// TIA Portal project "EbAndon v4_00_036" (V15) (continued)
   // pnText[239] := WSTRING#'//';
   // pnText[240] := WSTRING#'//';
   // pnText[241] := WSTRING#'//';
   // pnText[242] := WSTRING#'//';
   // pnText[243] := WSTRING#'//';
   // pnText[244] := WSTRING#'//';
   // pnText[245] := WSTRING#'//';
   // pnText[246] := WSTRING#'//';
   // pnText[247] := WSTRING#'//';
   // pnText[248] := WSTRING#'//';
   // pnText[249] := WSTRING#'//';
   // pnText[250] := WSTRING#'//';
   // pnText[251] := WSTRING#'//';
   // pnText[252] := WSTRING#'//';
   // pnText[253] := WSTRING#'//';
   // pnText[254] := WSTRING#'//';
   // pnText[255] := WSTRING#'//';
   // pnText[256] := WSTRING#'//';
   // pnText[257] := WSTRING#'//';
   // pnText[258] := WSTRING#'//';
   // pnText[259] := WSTRING#'//';
   // pnText[260] := WSTRING#'//';
   // pnText[261] := WSTRING#'//';
   // pnText[262] := WSTRING#'//';
   // pnText[263] := WSTRING#'//';
   // pnText[264] := WSTRING#'//';
   // pnText[265] := WSTRING#'//';
   // pnText[266] := WSTRING#'//';
   // pnText[267] := WSTRING#'//';
   // pnText[268] := WSTRING#'//';
   // pnText[269] := WSTRING#'//';
   // pnText[270] := WSTRING#'//';
   // pnText[271] := WSTRING#'//';
   // pnText[272] := WSTRING#'//';
   // pnText[273] := WSTRING#'//';
   // pnText[274] := WSTRING#'//';
   // pnText[275] := WSTRING#'//';
   // pnText[276] := WSTRING#'//';
   // pnText[277] := WSTRING#'//';
   // pnText[278] := WSTRING#'//';
   // pnText[279] := WSTRING#'//';
   // pnText[280] := WSTRING#'//';
   // pnText[281] := WSTRING#'//';
   // pnText[282] := WSTRING#'//';
   // pnText[283] := WSTRING#'//';
   // pnText[284] := WSTRING#'//';
   // pnText[285] := WSTRING#'//';
   // pnText[286] := WSTRING#'//';
   // pnText[287] := WSTRING#'//';
   // pnText[288] := WSTRING#'//';
   // pnText[289] := WSTRING#'//';
   // pnText[290] := WSTRING#'//';
   // pnText[291] := WSTRING#'//';
   // pnText[292] := WSTRING#'//';
   // pnText[293] := WSTRING#'//';
   // pnText[294] := WSTRING#'//';
   // pnText[295] := WSTRING#'//';
   // pnText[296] := WSTRING#'//';
   // pnText[297] := WSTRING#'//';
   // pnText[298] := WSTRING#'//';
   // pnText[299] := WSTRING#'//';
   // pnText[300] := WSTRING#'//';
   // pnText[301] := WSTRING#'//';
   // pnText[302] := WSTRING#'//';
   // pnText[303] := WSTRING#'//';
   // pnText[304] := WSTRING#'//';
   // pnText[305] := WSTRING#'//';
   // pnText[306] := WSTRING#'//';
   // pnText[307] := WSTRING#'//';
   // pnText[308] := WSTRING#'//';
   // pnText[309] := WSTRING#'//';
   // pnText[310] := WSTRING#'//';
   // pnText[311] := WSTRING#'//';
   // pnText[312] := WSTRING#'//';
   // pnText[313] := WSTRING#'//';
   // pnText[314] := WSTRING#'//';
   // pnText[315] := WSTRING#'//';
   // pnText[316] := WSTRING#'//';
   // pnText[317] := WSTRING#'//';
   // pnText[318] := WSTRING#'//';
   // pnText[319] := WSTRING#'//';
   // pnText[320] := WSTRING#'//';
   // pnText[321] := WSTRING#'//';
   // pnText[322] := WSTRING#'//';
   // pnText[323] := WSTRING#'//';
   // pnText[324] := WSTRING#'//';
   // pnText[325] := WSTRING#'//';
   // pnText[326] := WSTRING#'//';
   // pnText[327] := WSTRING#'//';
   // pnText[328] := WSTRING#'//';
   // pnText[329] := WSTRING#'//';
   // pnText[330] := WSTRING#'//';
   // pnText[331] := WSTRING#'//';
   // pnText[332] := WSTRING#'//';
   // pnText[333] := WSTRING#'//';
   // pnText[334] := WSTRING#'//';
   // pnText[335] := WSTRING#'//';
   // pnText[336] := WSTRING#'//';
   // pnText[337] := WSTRING#'//';
   // pnText[338] := WSTRING#'//';
   // pnText[339] := WSTRING#'//';
   // pnText[340] := WSTRING#'//';
   // pnText[341] := WSTRING#'//';
   // pnText[342] := WSTRING#'//';
   // pnText[343] := WSTRING#'//';
   // pnText[344] := WSTRING#'//';
   // pnText[345] := WSTRING#'//';
   // pnText[346] := WSTRING#'//';
   // pnText[347] := WSTRING#'//';
   // pnText[348] := WSTRING#'//';
   // pnText[349] := WSTRING#'//';
   // pnText[350] := WSTRING#'//';
   // pnText[351] := WSTRING#'//';
   // pnText[352] := WSTRING#'//';
   // pnText[353] := WSTRING#'//';
   // pnText[354] := WSTRING#'//';
   // pnText[355] := WSTRING#'//';
   // pnText[356] := WSTRING#'//';
   // pnText[357] := WSTRING#'//';
   // pnText[358] := WSTRING#'//';
   // pnText[359] := WSTRING#'//';
   // pnText[360] := WSTRING#'//';
   // pnText[361] := WSTRING#'//';
   // pnText[362] := WSTRING#'//';
   // pnText[363] := WSTRING#'//';
   // pnText[364] := WSTRING#'//';
   // pnText[365] := WSTRING#'//';
   // pnText[366] := WSTRING#'//';
   // pnText[367] := WSTRING#'//';
   // pnText[368] := WSTRING#'//';
   // pnText[369] := WSTRING#'//';
   // pnText[370] := WSTRING#'//';
   // pnText[371] := WSTRING#'//';
   // pnText[372] := WSTRING#'//';
   // pnText[373] := WSTRING#'//';
   // pnText[374] := WSTRING#'//';
   // pnText[375] := WSTRING#'//';
   // pnText[376] := WSTRING#'//';
   // pnText[377] := WSTRING#'//';
   // pnText[378] := WSTRING#'//';
   // pnText[379] := WSTRING#'//';
   // pnText[380] := WSTRING#'//';
   // pnText[381] := WSTRING#'//';
   // pnText[382] := WSTRING#'//';
   // pnText[383] := WSTRING#'//';
   // pnText[384] := WSTRING#'//';
   // pnText[385] := WSTRING#'//';
   // pnText[386] := WSTRING#'//';
   // pnText[387] := WSTRING#'//';
   // pnText[388] := WSTRING#'//';
   // pnText[389] := WSTRING#'//';
   // pnText[390] := WSTRING#'//';
   // pnText[391] := WSTRING#'//';
   // pnText[392] := WSTRING#'//';
   // pnText[393] := WSTRING#'//';
   // pnText[394] := WSTRING#'//';
   // pnText[395] := WSTRING#'//';
   // pnText[396] := WSTRING#'//';
   // pnText[397] := WSTRING#'//';
   // pnText[398] := WSTRING#'//';
   // pnText[399] := WSTRING#'//';
   // pnText[400] := WSTRING#'//';
   // pnText[401] := WSTRING#'//';
   // pnText[402] := WSTRING#'//';
   // pnText[403] := WSTRING#'//';
   // pnText[404] := WSTRING#'//';
   // pnText[405] := WSTRING#'//';
   // pnText[406] := WSTRING#'//';
   // pnText[407] := WSTRING#'//';
   // pnText[408] := WSTRING#'//';
   // pnText[409] := WSTRING#'//';
   // pnText[410] := WSTRING#'//';
   // pnText[411] := WSTRING#'//';
   // pnText[412] := WSTRING#'//';
   // pnText[413] := WSTRING#'//';
   // pnText[414] := WSTRING#'//';
   // pnText[415] := WSTRING#'//';
   // pnText[416] := WSTRING#'//';
   // pnText[417] := WSTRING#'//';
   // pnText[418] := WSTRING#'//';
   // pnText[419] := WSTRING#'//';
   // pnText[420] := WSTRING#'//';
   // pnText[421] := WSTRING#'//';
   // pnText[422] := WSTRING#'//';
   // pnText[423] := WSTRING#'//';
   // pnText[424] := WSTRING#'//';
   // pnText[425] := WSTRING#'//';
   // pnText[426] := WSTRING#'//';
   // pnText[427] := WSTRING#'//';
   // pnText[428] := WSTRING#'//';
   // pnText[429] := WSTRING#'//';
   // pnText[430] := WSTRING#'//';
   // pnText[431] := WSTRING#'//';
   // pnText[432] := WSTRING#'//';
   // pnText[433] := WSTRING#'//';
   // pnText[434] := WSTRING#'//';
   // pnText[435] := WSTRING#'//';
   // pnText[436] := WSTRING#'//';
   // pnText[437] := WSTRING#'//';
   // pnText[438] := WSTRING#'//';
   // pnText[439] := WSTRING#'//';
   // pnText[440] := WSTRING#'//';
   // pnText[441] := WSTRING#'//';
   // pnText[442] := WSTRING#'//';
   // pnText[443] := WSTRING#'//';
   // pnText[444] := WSTRING#'//';
   // pnText[445] := WSTRING#'//';
   // pnText[446] := WSTRING#'//';
   // pnText[447] := WSTRING#'//';
   // pnText[448] := WSTRING#'//';
   // pnText[449] := WSTRING#'//';
   // pnText[450] := WSTRING#'//';
   // pnText[451] := WSTRING#'//';
   // pnText[452] := WSTRING#'//';
   // pnText[453] := WSTRING#'//';
   // pnText[454] := WSTRING#'//';
   // pnText[455] := WSTRING#'//';
   // pnText[456] := WSTRING#'//';
   // pnText[457] := WSTRING#'//';
   // pnText[458] := WSTRING#'//';
   // pnText[459] := WSTRING#'//';
   // pnText[460] := WSTRING#'//';
   // pnText[461] := WSTRING#'//';
   // pnText[462] := WSTRING#'//';
   // pnText[463] := WSTRING#'//';
   // pnText[464] := WSTRING#'//';
   // pnText[465] := WSTRING#'//';
   // pnText[466] := WSTRING#'//';
   // pnText[467] := WSTRING#'//';
   // pnText[468] := WSTRING#'//';
   // pnText[469] := WSTRING#'//';
   // pnText[470] := WSTRING#'//';
   // pnText[471] := WSTRING#'//';
   // pnText[472] := WSTRING#'//';
   // pnText[473] := WSTRING#'//';
   // pnText[474] := WSTRING#'//';
   // pnText[475] := WSTRING#'//';
   // pnText[476] := WSTRING#'//';
   // pnText[477] := WSTRING#'//';
   // pnText[478] := WSTRING#'//';
   // pnText[479] := WSTRING#'//';
   // pnText[480] := WSTRING#'//';
   // pnText[481] := WSTRING#'//';
   // pnText[482] := WSTRING#'//';
   // pnText[483] := WSTRING#'//';
   // pnText[484] := WSTRING#'//';
   // pnText[485] := WSTRING#'//';
   // pnText[486] := WSTRING#'//';
   // pnText[487] := WSTRING#'//';
   // pnText[488] := WSTRING#'//';
   // pnText[489] := WSTRING#'//';
   // pnText[490] := WSTRING#'//';
   // pnText[491] := WSTRING#'//';
   // pnText[492] := WSTRING#'//';
   // pnText[493] := WSTRING#'//';
   // pnText[494] := WSTRING#'//';
   // pnText[495] := WSTRING#'//';
   // pnText[496] := WSTRING#'//';
   // pnText[497] := WSTRING#'//';
   // pnText[498] := WSTRING#'//';
   // pnText[499] := WSTRING#'//';
   // pnText[500] := WSTRING#'//';
   // pnText[501] := WSTRING#'//';
   // pnText[502] := WSTRING#'//';
   // pnText[503] := WSTRING#'//';
   // pnText[504] := WSTRING#'//';
   // pnText[505] := WSTRING#'//';
   // pnText[506] := WSTRING#'//';
   // pnText[507] := WSTRING#'//';
   // pnText[508] := WSTRING#'//';
   // pnText[509] := WSTRING#'//';
   // pnText[510] := WSTRING#'//';
   // pnText[511] := WSTRING#'//';
   // pnText[512] := WSTRING#'//';
   // pnText[513] := WSTRING#'//';
   // pnText[514] := WSTRING#'//';
   // pnText[515] := WSTRING#'//';
   // pnText[516] := WSTRING#'//';
   // pnText[517] := WSTRING#'//';
   // pnText[518] := WSTRING#'//';
   // pnText[519] := WSTRING#'//';
   // pnText[520] := WSTRING#'//';
   // pnText[521] := WSTRING#'//';
   // pnText[522] := WSTRING#'//';
   // pnText[523] := WSTRING#'//';
   // pnText[524] := WSTRING#'//';
   // pnText[525] := WSTRING#'//';
   // pnText[526] := WSTRING#'//';
   // pnText[527] := WSTRING#'//';
   // pnText[528] := WSTRING#'//';
   // pnText[529] := WSTRING#'//';
   // pnText[530] := WSTRING#'//';
   // pnText[531] := WSTRING#'//';
   // pnText[532] := WSTRING#'//';
   // pnText[533] := WSTRING#'//';
   // pnText[534] := WSTRING#'//';
   // pnText[535] := WSTRING#'//';
   // pnText[536] := WSTRING#'//';
   // pnText[537] := WSTRING#'//';
   // pnText[538] := WSTRING#'//';
   // pnText[539] := WSTRING#'//';
   // pnText[540] := WSTRING#'//';
   // pnText[541] := WSTRING#'//';
   // pnText[542] := WSTRING#'//';
   // pnText[543] := WSTRING#'//';
   // pnText[544] := WSTRING#'//';
   // pnText[545] := WSTRING#'//';
   // pnText[546] := WSTRING#'//';
   // pnText[547] := WSTRING#'//';
   // pnText[548] := WSTRING#'//';
   // pnText[549] := WSTRING#'//';
   // pnText[550] := WSTRING#'//';
   // pnText[551] := WSTRING#'//';
   // pnText[552] := WSTRING#'//';
   // pnText[553] := WSTRING#'//';
   // pnText[554] := WSTRING#'//';
   // pnText[555] := WSTRING#'//';
   // pnText[556] := WSTRING#'//';
   // pnText[557] := WSTRING#'//';
   // pnText[558] := WSTRING#'//';
   // pnText[559] := WSTRING#'//';
   // pnText[560] := WSTRING#'//';
   // pnText[561] := WSTRING#'//';
   // pnText[562] := WSTRING#'//';
   // pnText[563] := WSTRING#'//';
   // pnText[564] := WSTRING#'//';
   // pnText[565] := WSTRING#'//';
   // pnText[566] := WSTRING#'//';
   // pnText[567] := WSTRING#'//';
   // pnText[568] := WSTRING#'//';
   // pnText[569] := WSTRING#'//';
   // pnText[570] := WSTRING#'//';
   // pnText[571] := WSTRING#'//';
   // pnText[572] := WSTRING#'//';
   // pnText[573] := WSTRING#'//';
   // pnText[574] := WSTRING#'//';
   // pnText[575] := WSTRING#'//';
   // pnText[576] := WSTRING#'//';
   // pnText[577] := WSTRING#'//';
   // pnText[578] := WSTRING#'//';
   // pnText[579] := WSTRING#'//';
   // pnText[580] := WSTRING#'//';
   // pnText[581] := WSTRING#'//';
   // pnText[582] := WSTRING#'//';
   // pnText[583] := WSTRING#'//';
   // pnText[584] := WSTRING#'//';
   // pnText[585] := WSTRING#'//';
   // pnText[586] := WSTRING#'//';
   // pnText[587] := WSTRING#'//';
   // pnText[588] := WSTRING#'//';
   // pnText[589] := WSTRING#'//';
   // pnText[590] := WSTRING#'//';
   // pnText[591] := WSTRING#'//';
   // pnText[592] := WSTRING#'//';
   // pnText[593] := WSTRING#'//';
   // pnText[594] := WSTRING#'//';
   // pnText[595] := WSTRING#'//';
   // pnText[596] := WSTRING#'//';
   // pnText[597] := WSTRING#'//';
   // pnText[598] := WSTRING#'//';
   // pnText[599] := WSTRING#'//';
   // pnText[600] := WSTRING#'//';
   // pnText[601] := WSTRING#'//';
   // pnText[602] := WSTRING#'//';
   // pnText[603] := WSTRING#'//';
   // pnText[604] := WSTRING#'//';
   // pnText[605] := WSTRING#'//';
   // pnText[606] := WSTRING#'//';
   // pnText[607] := WSTRING#'//';
   // pnText[608] := WSTRING#'//';
   // pnText[609] := WSTRING#'//';
   // pnText[610] := WSTRING#'//';
   // pnText[611] := WSTRING#'//';
   // pnText[612] := WSTRING#'//';
   // pnText[613] := WSTRING#'//';
   // pnText[614] := WSTRING#'//';
   // pnText[615] := WSTRING#'//';
   // pnText[616] := WSTRING#'//';
   // pnText[617] := WSTRING#'//';
   // pnText[618] := WSTRING#'//';
   // pnText[619] := WSTRING#'//';
   // pnText[620] := WSTRING#'//';
   // pnText[621] := WSTRING#'//';
   // pnText[622] := WSTRING#'//';
   // pnText[623] := WSTRING#'//';
   // pnText[624] := WSTRING#'//';
   // pnText[625] := WSTRING#'//';
   // pnText[626] := WSTRING#'//';
   // pnText[627] := WSTRING#'//';
   // pnText[628] := WSTRING#'//';
   // pnText[629] := WSTRING#'//';
   // pnText[630] := WSTRING#'//';
   // pnText[631] := WSTRING#'//';
   // pnText[632] := WSTRING#'//';
   // pnText[633] := WSTRING#'//';
   // pnText[634] := WSTRING#'//';
   // pnText[635] := WSTRING#'//';
   // pnText[636] := WSTRING#'//';
   // pnText[637] := WSTRING#'//';
   // pnText[638] := WSTRING#'//';
   // pnText[639] := WSTRING#'//';
   // pnText[640] := WSTRING#'//';
   // pnText[641] := WSTRING#'//';
   // pnText[642] := WSTRING#'//';
   // pnText[643] := WSTRING#'//';
   // pnText[644] := WSTRING#'//';
   // pnText[645] := WSTRING#'//';
   // pnText[646] := WSTRING#'//';
   // pnText[647] := WSTRING#'//';
   // pnText[648] := WSTRING#'//';
   // pnText[649] := WSTRING#'//';
   // pnText[650] := WSTRING#'//';
   // pnText[651] := WSTRING#'//';
   // pnText[652] := WSTRING#'//';
   // pnText[653] := WSTRING#'//';
   // pnText[654] := WSTRING#'//';
   // pnText[655] := WSTRING#'//';
   // pnText[656] := WSTRING#'//';
   // pnText[657] := WSTRING#'//';
   // pnText[658] := WSTRING#'//';
   // pnText[659] := WSTRING#'//';
   // pnText[660] := WSTRING#'//';
   // pnText[661] := WSTRING#'//';
   // pnText[662] := WSTRING#'//';
   // pnText[663] := WSTRING#'//';
   // pnText[664] := WSTRING#'//';
   // pnText[665] := WSTRING#'//';
   // pnText[666] := WSTRING#'//';
   // pnText[667] := WSTRING#'//';
   // pnText[668] := WSTRING#'//';
   // pnText[669] := WSTRING#'//';
   // pnText[670] := WSTRING#'//';
   // pnText[671] := WSTRING#'//';
   // pnText[672] := WSTRING#'//';
   // pnText[673] := WSTRING#'//';
   // pnText[674] := WSTRING#'//';
   // pnText[675] := WSTRING#'//';
   // pnText[676] := WSTRING#'//';
   // pnText[677] := WSTRING#'//';
   // pnText[678] := WSTRING#'//';
   // pnText[679] := WSTRING#'//';
   // pnText[680] := WSTRING#'//';
   // pnText[681] := WSTRING#'//';
   // pnText[682] := WSTRING#'//';
   // pnText[683] := WSTRING#'//';
   // pnText[684] := WSTRING#'//';
   // pnText[685] := WSTRING#'//';
   // pnText[686] := WSTRING#'//';
   // pnText[687] := WSTRING#'//';
   // pnText[688] := WSTRING#'//';
   // pnText[689] := WSTRING#'//';
   // pnText[690] := WSTRING#'//';
   // pnText[691] := WSTRING#'//';
   // pnText[692] := WSTRING#'//';
   // pnText[693] := WSTRING#'//';
   // pnText[694] := WSTRING#'//';
   // pnText[695] := WSTRING#'//';
   // pnText[696] := WSTRING#'//';
   // pnText[697] := WSTRING#'//';
   // pnText[698] := WSTRING#'//';
   // pnText[699] := WSTRING#'//';
   // pnText[700] := WSTRING#'//';
   // pnText[701] := WSTRING#'//';
   // pnText[702] := WSTRING#'//';
   // pnText[703] := WSTRING#'//';
   // pnText[704] := WSTRING#'//';
   // pnText[705] := WSTRING#'//';
   // pnText[706] := WSTRING#'//';
   // pnText[707] := WSTRING#'//';
   // pnText[708] := WSTRING#'//';
   // pnText[709] := WSTRING#'//';
   // pnText[710] := WSTRING#'//';
   // pnText[711] := WSTRING#'//';
   // pnText[712] := WSTRING#'//';
   // pnText[713] := WSTRING#'//';
   // pnText[714] := WSTRING#'//';
   // pnText[715] := WSTRING#'//';
   // pnText[716] := WSTRING#'//';
   // pnText[717] := WSTRING#'//';
   // pnText[718] := WSTRING#'//';
   // pnText[719] := WSTRING#'//';
   // pnText[720] := WSTRING#'//';
   // pnText[721] := WSTRING#'//';
   // pnText[722] := WSTRING#'//';
   // pnText[723] := WSTRING#'//';
   // pnText[724] := WSTRING#'//';
   // pnText[725] := WSTRING#'//';
   // pnText[726] := WSTRING#'//';
   // pnText[727] := WSTRING#'//';
   // pnText[728] := WSTRING#'//';
   // pnText[729] := WSTRING#'//';
   // pnText[730] := WSTRING#'//';
   // pnText[731] := WSTRING#'//';
   // pnText[732] := WSTRING#'//';
   // pnText[733] := WSTRING#'//';
   // pnText[734] := WSTRING#'//';
   // pnText[735] := WSTRING#'//';
   // pnText[736] := WSTRING#'//';
   // pnText[737] := WSTRING#'//';
   // pnText[738] := WSTRING#'//';
   // pnText[739] := WSTRING#'//';
   // pnText[740] := WSTRING#'//';
   // pnText[741] := WSTRING#'//';
   // pnText[742] := WSTRING#'//';
   // pnText[743] := WSTRING#'//';
   // pnText[744] := WSTRING#'//';
   // pnText[745] := WSTRING#'//';
   // pnText[746] := WSTRING#'//';
   // pnText[747] := WSTRING#'//';
   // pnText[748] := WSTRING#'//';
   // pnText[749] := WSTRING#'//';
   // pnText[750] := WSTRING#'//';
   // pnText[751] := WSTRING#'//';
   // pnText[752] := WSTRING#'//';
   // pnText[753] := WSTRING#'//';
   // pnText[754] := WSTRING#'//';
   // pnText[755] := WSTRING#'//';
   // pnText[756] := WSTRING#'//';
   // pnText[757] := WSTRING#'//';
   // pnText[758] := WSTRING#'//';
   // pnText[759] := WSTRING#'//';
   // pnText[760] := WSTRING#'//';
   // pnText[761] := WSTRING#'//';
   // pnText[762] := WSTRING#'//';
   // pnText[763] := WSTRING#'//';
   // pnText[764] := WSTRING#'//';
   // pnText[765] := WSTRING#'//';
   // pnText[766] := WSTRING#'//';
   // pnText[767] := WSTRING#'//';
   // pnText[768] := WSTRING#'//';
   // pnText[769] := WSTRING#'//';
   // pnText[770] := WSTRING#'//';
   // pnText[771] := WSTRING#'//';
   // pnText[772] := WSTRING#'//';
   // pnText[773] := WSTRING#'//';
   // pnText[774] := WSTRING#'//';
   // pnText[775] := WSTRING#'//';
   // pnText[776] := WSTRING#'//';
   // pnText[777] := WSTRING#'//';
   // pnText[778] := WSTRING#'//';
   // pnText[779] := WSTRING#'//';
   // pnText[780] := WSTRING#'//';
   // pnText[781] := WSTRING#'//';
   // pnText[782] := WSTRING#'//';
   // pnText[783] := WSTRING#'//';
   // pnText[784] := WSTRING#'//';
   // pnText[785] := WSTRING#'//';
   // pnText[786] := WSTRING#'//';
   // pnText[787] := WSTRING#'//';
   // pnText[788] := WSTRING#'//';
   // pnText[789] := WSTRING#'//';
   // pnText[790] := WSTRING#'//';
   // pnText[791] := WSTRING#'//';
   // pnText[792] := WSTRING#'//';
   // pnText[793] := WSTRING#'//';
   // pnText[794] := WSTRING#'//';
   // pnText[795] := WSTRING#'//';
   // pnText[796] := WSTRING#'//';
   // pnText[797] := WSTRING#'//';
   // pnText[798] := WSTRING#'//';
   // pnText[799] := WSTRING#'//';
   // pnText[800] := WSTRING#'//';
   // pnText[801] := WSTRING#'//';
   // pnText[802] := WSTRING#'//';
   // pnText[803] := WSTRING#'//';
   // pnText[804] := WSTRING#'//';
   // pnText[805] := WSTRING#'//';
   // pnText[806] := WSTRING#'//';
   // pnText[807] := WSTRING#'//';
   // pnText[808] := WSTRING#'//';
   // pnText[809] := WSTRING#'//';
   // pnText[810] := WSTRING#'//';
   // pnText[811] := WSTRING#'//';
   // pnText[812] := WSTRING#'//';
   // pnText[813] := WSTRING#'//';
   // pnText[814] := WSTRING#'//';
   // pnText[815] := WSTRING#'//';
   // pnText[816] := WSTRING#'//';
   // pnText[817] := WSTRING#'//';
   // pnText[818] := WSTRING#'//';
   // pnText[819] := WSTRING#'//';
   // pnText[820] := WSTRING#'//';
   // pnText[821] := WSTRING#'//';
   // pnText[822] := WSTRING#'//';
   // pnText[823] := WSTRING#'//';
   // pnText[824] := WSTRING#'//';
   // pnText[825] := WSTRING#'//';
   // pnText[826] := WSTRING#'//';
   // pnText[827] := WSTRING#'//';
   // pnText[828] := WSTRING#'//';
   // pnText[829] := WSTRING#'//';
   // pnText[830] := WSTRING#'//';
   // pnText[831] := WSTRING#'//';
   // pnText[832] := WSTRING#'//';
   // pnText[833] := WSTRING#'//';
   // pnText[834] := WSTRING#'//';
   // pnText[835] := WSTRING#'//';
   // pnText[836] := WSTRING#'//';
   // pnText[837] := WSTRING#'//';
   // pnText[838] := WSTRING#'//';
   // pnText[839] := WSTRING#'//';
   // pnText[840] := WSTRING#'//';
   // pnText[841] := WSTRING#'//';
   // pnText[842] := WSTRING#'//';
   // pnText[843] := WSTRING#'//';
   // pnText[844] := WSTRING#'//';
   // pnText[845] := WSTRING#'//';
   // pnText[846] := WSTRING#'//';
   // pnText[847] := WSTRING#'//';
   // pnText[848] := WSTRING#'//';
   // pnText[849] := WSTRING#'//';
   // pnText[850] := WSTRING#'//';
   // pnText[851] := WSTRING#'//';
   // pnText[852] := WSTRING#'//';
   // pnText[853] := WSTRING#'//';
   // pnText[854] := WSTRING#'//';
   // pnText[855] := WSTRING#'//';
   // pnText[856] := WSTRING#'//';
   // pnText[857] := WSTRING#'//';
   // pnText[858] := WSTRING#'//';
   // pnText[859] := WSTRING#'//';
   // pnText[860] := WSTRING#'//';
   // pnText[861] := WSTRING#'//';
   // pnText[862] := WSTRING#'//';
   // pnText[863] := WSTRING#'//';
   // pnText[864] := WSTRING#'//';
   // pnText[865] := WSTRING#'//';
   // pnText[866] := WSTRING#'//';
   // pnText[867] := WSTRING#'//';
   // pnText[868] := WSTRING#'//';
   // pnText[869] := WSTRING#'//';
   // pnText[870] := WSTRING#'//';
   // pnText[871] := WSTRING#'//';
   // pnText[872] := WSTRING#'//';
   // pnText[873] := WSTRING#'//';
   // pnText[874] := WSTRING#'//';
   // pnText[875] := WSTRING#'//';
   // pnText[876] := WSTRING#'//';
   // pnText[877] := WSTRING#'//';
   // pnText[878] := WSTRING#'//';
   // pnText[879] := WSTRING#'//';
   // pnText[880] := WSTRING#'//';
   // pnText[881] := WSTRING#'//';
   // pnText[882] := WSTRING#'//';
   // pnText[883] := WSTRING#'//';
   // pnText[884] := WSTRING#'//';
   // pnText[885] := WSTRING#'//';
   // pnText[886] := WSTRING#'//';
   // pnText[887] := WSTRING#'//';
   // pnText[888] := WSTRING#'//';
   // pnText[889] := WSTRING#'//';
   // pnText[890] := WSTRING#'//';
   // pnText[891] := WSTRING#'//';
   // pnText[892] := WSTRING#'//';
   // pnText[893] := WSTRING#'//';
   // pnText[894] := WSTRING#'//';
   // pnText[895] := WSTRING#'//';
   // pnText[896] := WSTRING#'//';
   // pnText[897] := WSTRING#'//';
   // pnText[898] := WSTRING#'//';
   // pnText[899] := WSTRING#'//';
   // pnText[900] := WSTRING#'//';
   // pnText[901] := WSTRING#'//';
   // pnText[902] := WSTRING#'//';
   // pnText[903] := WSTRING#'//';
   // pnText[904] := WSTRING#'//';
   // pnText[905] := WSTRING#'//';
   // pnText[906] := WSTRING#'//';
   // pnText[907] := WSTRING#'//';
   // pnText[908] := WSTRING#'//';
   // pnText[909] := WSTRING#'//';
   // pnText[910] := WSTRING#'//';
   // pnText[911] := WSTRING#'//';
   // pnText[912] := WSTRING#'//';
   // pnText[913] := WSTRING#'//';
   // pnText[914] := WSTRING#'//';
   // pnText[915] := WSTRING#'//';
   // pnText[916] := WSTRING#'//';
   // pnText[917] := WSTRING#'//';
   // pnText[918] := WSTRING#'//';
   // pnText[919] := WSTRING#'//';
   // pnText[920] := WSTRING#'//';
   // pnText[921] := WSTRING#'//';
   // pnText[922] := WSTRING#'//';
   // pnText[923] := WSTRING#'//';
   // pnText[924] := WSTRING#'//';
   // pnText[925] := WSTRING#'//';
   // pnText[926] := WSTRING#'//';
   // pnText[927] := WSTRING#'//';
   // pnText[928] := WSTRING#'//';
   // pnText[929] := WSTRING#'//';
   // pnText[930] := WSTRING#'//';
   // pnText[931] := WSTRING#'//';
   // pnText[932] := WSTRING#'//';
   // pnText[933] := WSTRING#'//';
   // pnText[934] := WSTRING#'//';
   // pnText[935] := WSTRING#'//';
   // pnText[936] := WSTRING#'//';
   // pnText[937] := WSTRING#'//';
   // pnText[938] := WSTRING#'//';
   // pnText[939] := WSTRING#'//';
   // pnText[940] := WSTRING#'//';
   // pnText[941] := WSTRING#'//';
   // pnText[942] := WSTRING#'//';
   // pnText[943] := WSTRING#'//';
   // pnText[944] := WSTRING#'//';
   // pnText[945] := WSTRING#'//';
   // pnText[946] := WSTRING#'//';
   // pnText[947] := WSTRING#'//';
   // pnText[948] := WSTRING#'//';
   // pnText[949] := WSTRING#'//';
   // pnText[950] := WSTRING#'//';
   // pnText[951] := WSTRING#'//';
   // pnText[952] := WSTRING#'//';
   // pnText[953] := WSTRING#'//';
   // pnText[954] := WSTRING#'//';
   // pnText[955] := WSTRING#'//';
   // pnText[956] := WSTRING#'//';
   // pnText[957] := WSTRING#'//';
   // pnText[958] := WSTRING#'//';
   // pnText[959] := WSTRING#'//';
   // pnText[960] := WSTRING#'//';
   // pnText[961] := WSTRING#'//';
   // pnText[962] := WSTRING#'//';
   // pnText[963] := WSTRING#'//';
   // pnText[964] := WSTRING#'//';
   // pnText[965] := WSTRING#'//';
   // pnText[966] := WSTRING#'//';
   // pnText[967] := WSTRING#'//';
   // pnText[968] := WSTRING#'//';
   // pnText[969] := WSTRING#'//';
   // pnText[970] := WSTRING#'//';
   // pnText[971] := WSTRING#'//';
   // pnText[972] := WSTRING#'//';
   // pnText[973] := WSTRING#'//';
   // pnText[974] := WSTRING#'//';
   // pnText[975] := WSTRING#'//';
   // pnText[976] := WSTRING#'//';
   // pnText[977] := WSTRING#'//';
   // pnText[978] := WSTRING#'//';
   // pnText[979] := WSTRING#'//';
   // pnText[980] := WSTRING#'//';
   // pnText[981] := WSTRING#'//';
   // pnText[982] := WSTRING#'//';
   // pnText[983] := WSTRING#'//';
   // pnText[984] := WSTRING#'//';
   // pnText[985] := WSTRING#'//';
   // pnText[986] := WSTRING#'//';
   // pnText[987] := WSTRING#'//';
   // pnText[988] := WSTRING#'//';
   // pnText[989] := WSTRING#'//';
   // pnText[990] := WSTRING#'//';
   // pnText[991] := WSTRING#'//';
   // pnText[992] := WSTRING#'//';
   // pnText[993] := WSTRING#'//';
   // pnText[994] := WSTRING#'//';
   // pnText[995] := WSTRING#'//';
   // pnText[996] := WSTRING#'//';
   // pnText[997] := WSTRING#'//';
   // pnText[998] := WSTRING#'//';
   // pnText[999] := WSTRING#'//';
END_TYPE

TYPE "Selected Wips"
   STRUCT
      count : Int;
      wips : Array[0.."WIP_COUNT"] of DInt;
   END_STRUCT;
END_TYPE

TYPE "Selected Buttons"
   STRUCT
      btns : Array[0.."BUTTON_COUNT"] of Bool;
      count : Int;
   END_STRUCT;
END_TYPE

TYPE "Setting Meta Data"
   STRUCT
      selectable_stations : "Selectable Stations";
      selectable_wips : "Selectable Wips";
      selected_btns : "Selected Buttons";
      selected_stations : "Selected Stations";
      selected_wips : "Selected Wips";
      station_selection_change : "Station Selection Change";
      button_selection_change : "Selected_Buttons.Selection_Change.UDT";
   END_STRUCT;
END_TYPE

TYPE "Nav Bar Data"
   STRUCT
      hmi : "Nav Bar Data: HMI";
      plc : "Nav Bar Data: PLC";
   END_STRUCT;
END_TYPE

TYPE "Intersecting WIPs Arrays"
   STRUCT
      count : Int;
      WIPS_intersection : Array[0.."WIP_COUNT"] of DInt;
   END_STRUCT;
END_TYPE

TYPE "Initialize Excel Data: States"
   STRUCT
      active_wip_to_hmi_station_list : Bool;
      active_wip_to_master_station_list : Bool;
      pn_code_to_kp8_station : Bool;
      pn_code_to_saved_wips : Bool;
      wip_code_to_saved_wips : Bool;
   END_STRUCT;
END_TYPE

TYPE "Push Button Data: State Change Data"
   STRUCT
      actuate : "State Changes: Bool";
      animate : "State Changes: USInt";
      enable : "State Changes: Bool";
      label : "State Changes: WString";
      listSelect : "State Changes: UInt";
      visible : "State Changes: Bool";
   END_STRUCT;
END_TYPE

TYPE "IO Field: State Change Data"
   STRUCT
      animate : "State Changes: USInt";
      enable : "State Changes: Bool";
      input_finished : "State Changes: Bool";
      value : "State Changes: WString";
      visible : "State Changes: Bool";
   END_STRUCT;
END_TYPE

TYPE "Part_Number_Double.UDT"
   STRUCT
      single_actuate : Bool;
      single_animate : USInt;
      single_enable : Bool;
      single_input_finished : Bool;
      single_value : WString[40];
      single_visible : Bool;
      double_actuate : Bool;
      double_animate : USInt;
      double_enable : Bool;
      double_input_finished_top : Bool;
      double_input_finished_bottom : Bool;
      double_value_top : WString[40];
      double_value_bottom : WString[40];
      double_visible : Bool;
   END_STRUCT;
END_TYPE

TYPE "Selected_WIP_Table.Selected_Element"
   STRUCT
      station_pointer : Int;
      wip_pointer : DInt;
   END_STRUCT;
END_TYPE

TYPE "Selected_WIP_Table.Selected_Array"
   STRUCT
      me : Array[0..99] of "Selected_WIP_Table.Selected_Element";
   END_STRUCT;
END_TYPE

TYPE "Part_Number_Double.State_Change.UDT"
   STRUCT
      single : Struct
         actuate : "State Changes: Bool";
         animate : "State Changes: USInt";
         enable : "State Changes: Bool";
         input_finished : "State Changes: Bool";
         value : "State Changes: WString";
         visible : "State Changes: Bool";
      END_STRUCT;
      double : Struct
         actuate : "State Changes: Bool";
         animate : "State Changes: USInt";
         enable : "State Changes: Bool";
         visible : "State Changes: Bool";
         top : Struct
            input_finished : "State Changes: Bool";
            value : "State Changes: WString";
         END_STRUCT;
         bottom : Struct
            input_finished : "State Changes: Bool";
            value : "State Changes: WString";
         END_STRUCT;
      END_STRUCT;
   END_STRUCT;
END_TYPE

TYPE "Selected_Buttons.Selection_Change.UDT"
   STRUCT
      falling : Bool;
      rising : Bool;
      selection_change : Bool;
      button_index : Int := -1;
   END_STRUCT;
END_TYPE

// folder: From Excel

TYPE "From Excel: Codes Single Wip"
VERSION : 0.1
   STRUCT
      pStn : Int := -1;
      pnCode : Array[0.."BUTTON_COUNT"] of DInt;
   END_STRUCT;
END_TYPE

TYPE "From Excel: Codes Multiple Wips"
VERSION : 0.1
   STRUCT
      pStn : Int := -1;
      wip : Array[0.."WIP_COUNT"] of Struct
         wipCode : DInt;
         pnCode : Array[0.."BUTTON_COUNT"] of DInt;
      END_STRUCT;
   END_STRUCT;
END_TYPE

